screen "101_SDC_PN_Diag128_255" 1280x800, template "SDC"
   on GenerateScreen: SetTag("_intern_BILD_Nr", 101); SetTag("PN_PB\PN\IOSys_ID", 100)
   on ClearScreen: SetTag("_intern_BILD_Nr", 0)
   TextField "OBJECT_674" at 262,49 size 227x27; Text 'ProfiNet-System'
      Visibility <- "PN_PB\IO_Sys_ID"
   Button "Schaltfläche_2" at 240,609 size 107x60; TextOff 'Diagnose PN 101'
      on Press: SetTag("PN_PB\PN\IOSys_ID", 101)
      Visibility <- "PN_PB\IO_Sys_ID"
   Button "Schaltfläche_1" at 240,609 size 107x60; TextOff 'Diagnose PN 100'
      on Press: SetTag("PN_PB\PN\IOSys_ID", 100)
      Visibility <- "PN_PB\IO_Sys_ID"
   Button "Schaltfläche_4" at 573,45 size 359x37; TextOff 'ProfiNet-Teilnehmer 0 - 127'
      on Release: ActivateScreen("100_SDC_PN_Diag0_127", 0)
   GraphicView "OBJECT_496" at 1179,498 size 60x43; Picture "PB_Array_blau_3"
   TextField "OBJECT_497" at 1189,510 size 40x20; Text '1'
   GraphicView "OBJECT_498" at 1179,545 size 60x43; Picture "PB_Array_grün_3"
   TextField "OBJECT_499" at 1189,556 size 40x20; Text '1'
   TextField "OBJECT_500" at 1189,600 size 40x20; Text '1'
   GraphicView "OBJECT_501" at 1179,590 size 60x43; Picture "PB_Array_grün_3"
   TextField "OBJECT_502" at 1189,600 size 40x20; Text '1'
   TextField "OBJECT_504" at 922,505 size 257x31; Text 'Teilnehmer nicht vorhanden'
   TextField "OBJECT_505" at 922,597 size 193x33; Text 'Teilnehmer gestört'
   TextField "OBJECT_506" at 922,552 size 213x33; Text 'Teilnehmer vorhanden'
   TextField "OBJECT_670" at 902,469 size 111x35; Text 'Legende:'
   IOField "OBJECT_675" at 497,50 size 47x29; FormatPattern 999
      ProcessValue <- "PN_PB\IO_Sys_ID"
   TextField "OBJECT_513" at 255,503 size 104x29; Text 'Ort:'
   TextField "OBJECT_514" at 255,533 size 104x31; Text 'Typ:'
   TextField "OBJECT_515" at 255,563 size 131x29; Text 'Bezeichnung:'
   IOField "OBJECT_516" at 399,503 size 167x29; FormatPattern ????????????
      ProcessValue <- "PN_PB\Teiln_Nr_Ort"
   IOField "OBJECT_517" at 399,533 size 156x31; FormatPattern ????????????
      ProcessValue <- "PN_PB\Teiln_Nr_Typ"
   IOField "OBJECT_518" at 399,563 size 253x29; FormatPattern ????????????????????
      ProcessValue <- "PN_PB\Teiln_Nr_Bez"
   IOField "OBJECT_658" at 483,473 size 57x27; FormatPattern 999
      ProcessValue <- "PN_PB\PN\Teiln_Nr"
      Appearance <- "Trigger"
   TextField "OBJECT_679" at 587,473 size 67x25; Text 'Trigger'
      Appearance <- "Trigger"
   GraphicIOField "OBJECT_16" at 749,88 size 60x43; PictureList "PB_Slave_Bit15_3"
      ProcessValue <- "PN_PB\PTMUX_P_TLN129_144"
   GraphicIOField "OBJECT_151" at 813,88 size 60x43; PictureList "PB_Slave_Bit14_3"
      ProcessValue <- "PN_PB\PTMUX_P_TLN129_144"
   GraphicIOField "OBJECT_967" at 874,409 size 60x43; PictureList "PB_Slave_Bit13_3"
      ProcessValue <- "PN_PB\PTMUX_P_TLN241_256"
   GraphicIOField "OBJECT_968" at 1062,409 size 60x43; PictureList "PB_Slave_Bit10_3"
      ProcessValue <- "PN_PB\PTMUX_P_TLN241_256"
   GraphicIOField "OBJECT_969" at 1125,409 size 60x43; PictureList "PB_Slave_Bit9_3"
      ProcessValue <- "PN_PB\PTMUX_P_TLN241_256"
   GraphicIOField "OBJECT_970" at 1187,409 size 60x43; PictureList "PB_Slave_Bit8_3"
      ProcessValue <- "PN_PB\PTMUX_P_TLN241_256"
   GraphicIOField "OBJECT_971" at 999,409 size 60x43; PictureList "PB_Slave_Bit11_3"
      ProcessValue <- "PN_PB\PTMUX_P_TLN241_256"
   GraphicIOField "OBJECT_972" at 811,409 size 60x43; PictureList "PB_Slave_Bit14_3"
      ProcessValue <- "PN_PB\PTMUX_P_TLN241_256"
   GraphicIOField "OBJECT_973" at 937,409 size 60x43; PictureList "PB_Slave_Bit12_3"
      ProcessValue <- "PN_PB\PTMUX_P_TLN241_256"
   GraphicIOField "OBJECT_974" at 749,409 size 60x43; PictureList "PB_Slave_Bit15_3"
      ProcessValue <- "PN_PB\PTMUX_P_TLN241_256"
   GraphicIOField "OBJECT_1030" at 310,409 size 60x43; PictureList "PB_Slave_Bit6_3"
      ProcessValue <- "PN_PB\PTMUX_P_TLN241_256"
   GraphicIOField "OBJECT_1031" at 373,409 size 60x43; PictureList "PB_Slave_Bit5_3"
      ProcessValue <- "PN_PB\PTMUX_P_TLN241_256"
   GraphicIOField "OBJECT_1032" at 435,409 size 60x43; PictureList "PB_Slave_Bit4_3"
      ProcessValue <- "PN_PB\PTMUX_P_TLN241_256"
   GraphicIOField "OBJECT_1033" at 561,409 size 60x43; PictureList "PB_Slave_Bit2_3"
      ProcessValue <- "PN_PB\PTMUX_P_TLN241_256"
   GraphicIOField "OBJECT_1034" at 623,409 size 60x43; PictureList "PB_Slave_Bit1_3"
      ProcessValue <- "PN_PB\PTMUX_P_TLN241_256"
   GraphicIOField "OBJECT_1035" at 686,409 size 60x43; PictureList "PB_Slave_Bit0_3"
      ProcessValue <- "PN_PB\PTMUX_P_TLN241_256"
   GraphicIOField "OBJECT_1036" at 498,409 size 60x43; PictureList "PB_Slave_Bit3_3"
      ProcessValue <- "PN_PB\PTMUX_P_TLN241_256"
   GraphicIOField "OBJECT_1037" at 247,409 size 60x43; PictureList "PB_Slave_Bit7_3"
      ProcessValue <- "PN_PB\PTMUX_P_TLN241_256"
   GraphicIOField "OBJECT_983" at 310,133 size 60x43; PictureList "PB_Slave_Bit6_3"
      ProcessValue <- "PN_PB\PTMUX_P_TLN145_160"
   GraphicIOField "OBJECT_12" at 937,88 size 60x43; PictureList "PB_Slave_Bit12_3"
      ProcessValue <- "PN_PB\PTMUX_P_TLN129_144"
   GraphicIOField "OBJECT_13" at 310,88 size 60x43; PictureList "PB_Slave_Bit6_3"
      ProcessValue <- "PN_PB\PTMUX_P_TLN129_144"
   GraphicIOField "OBJECT_213" at 1062,88 size 60x43; PictureList "PB_Slave_Bit10_3"
      ProcessValue <- "PN_PB\PTMUX_P_TLN129_144"
   GraphicIOField "OBJECT_916" at 1125,88 size 60x43; PictureList "PB_Slave_Bit9_3"
      ProcessValue <- "PN_PB\PTMUX_P_TLN129_144"
   GraphicIOField "OBJECT_917" at 1187,88 size 60x43; PictureList "PB_Slave_Bit8_3"
      ProcessValue <- "PN_PB\PTMUX_P_TLN129_144"
   GraphicIOField "OBJECT_918" at 999,88 size 60x43; PictureList "PB_Slave_Bit11_3"
      ProcessValue <- "PN_PB\PTMUX_P_TLN129_144"
   GraphicIOField "OBJECT_919" at 749,133 size 60x43; PictureList "PB_Slave_Bit15_3"
      ProcessValue <- "PN_PB\PTMUX_P_TLN145_160"
   GraphicIOField "OBJECT_920" at 811,133 size 60x43; PictureList "PB_Slave_Bit14_3"
      ProcessValue <- "PN_PB\PTMUX_P_TLN145_160"
   GraphicIOField "OBJECT_921" at 874,133 size 60x43; PictureList "PB_Slave_Bit13_3"
      ProcessValue <- "PN_PB\PTMUX_P_TLN145_160"
   GraphicIOField "OBJECT_922" at 937,133 size 60x43; PictureList "PB_Slave_Bit12_3"
      ProcessValue <- "PN_PB\PTMUX_P_TLN145_160"
   GraphicIOField "OBJECT_923" at 1062,133 size 60x43; PictureList "PB_Slave_Bit10_3"
      ProcessValue <- "PN_PB\PTMUX_P_TLN145_160"
   GraphicIOField "OBJECT_924" at 1125,133 size 60x43; PictureList "PB_Slave_Bit9_3"
      ProcessValue <- "PN_PB\PTMUX_P_TLN145_160"
   GraphicIOField "OBJECT_925" at 1187,133 size 60x43; PictureList "PB_Slave_Bit8_3"
      ProcessValue <- "PN_PB\PTMUX_P_TLN145_160"
   GraphicIOField "OBJECT_926" at 999,133 size 60x43; PictureList "PB_Slave_Bit11_3"
      ProcessValue <- "PN_PB\PTMUX_P_TLN145_160"
   GraphicIOField "OBJECT_927" at 749,179 size 60x43; PictureList "PB_Slave_Bit15_3"
      ProcessValue <- "PN_PB\PTMUX_P_TLN161_176"
   GraphicIOField "OBJECT_928" at 874,179 size 60x43; PictureList "PB_Slave_Bit13_3"
      ProcessValue <- "PN_PB\PTMUX_P_TLN161_176"
   GraphicIOField "OBJECT_929" at 937,179 size 60x43; PictureList "PB_Slave_Bit12_3"
      ProcessValue <- "PN_PB\PTMUX_P_TLN161_176"
   GraphicIOField "OBJECT_930" at 1062,179 size 60x43; PictureList "PB_Slave_Bit10_3"
      ProcessValue <- "PN_PB\PTMUX_P_TLN161_176"
   GraphicIOField "OBJECT_931" at 1125,179 size 60x43; PictureList "PB_Slave_Bit9_3"
      ProcessValue <- "PN_PB\PTMUX_P_TLN161_176"
   GraphicIOField "OBJECT_932" at 1187,179 size 60x43; PictureList "PB_Slave_Bit8_3"
      ProcessValue <- "PN_PB\PTMUX_P_TLN161_176"
   GraphicIOField "OBJECT_933" at 999,179 size 60x43; PictureList "PB_Slave_Bit11_3"
      ProcessValue <- "PN_PB\PTMUX_P_TLN161_176"
   GraphicIOField "OBJECT_934" at 811,179 size 60x43; PictureList "PB_Slave_Bit14_3"
      ProcessValue <- "PN_PB\PTMUX_P_TLN161_176"
   GraphicIOField "OBJECT_935" at 749,224 size 60x43; PictureList "PB_Slave_Bit15_3"
      ProcessValue <- "PN_PB\PTMUX_P_TLN177_192"
   GraphicIOField "OBJECT_936" at 874,224 size 60x43; PictureList "PB_Slave_Bit13_3"
      ProcessValue <- "PN_PB\PTMUX_P_TLN177_192"
   GraphicIOField "OBJECT_937" at 937,224 size 60x43; PictureList "PB_Slave_Bit12_3"
      ProcessValue <- "PN_PB\PTMUX_P_TLN177_192"
   GraphicIOField "OBJECT_938" at 1062,224 size 60x43; PictureList "PB_Slave_Bit10_3"
      ProcessValue <- "PN_PB\PTMUX_P_TLN177_192"
   GraphicIOField "OBJECT_939" at 1125,224 size 60x43; PictureList "PB_Slave_Bit9_3"
      ProcessValue <- "PN_PB\PTMUX_P_TLN177_192"
   GraphicIOField "OBJECT_940" at 1187,224 size 60x43; PictureList "PB_Slave_Bit8_3"
      ProcessValue <- "PN_PB\PTMUX_P_TLN177_192"
   GraphicIOField "OBJECT_941" at 999,224 size 60x43; PictureList "PB_Slave_Bit11_3"
      ProcessValue <- "PN_PB\PTMUX_P_TLN177_192"
   GraphicIOField "OBJECT_942" at 811,224 size 60x43; PictureList "PB_Slave_Bit14_3"
      ProcessValue <- "PN_PB\PTMUX_P_TLN177_192"
   GraphicIOField "OBJECT_943" at 749,269 size 60x43; PictureList "PB_Slave_Bit15_3"
      ProcessValue <- "PN_PB\PTMUX_P_TLN193_208"
   GraphicIOField "OBJECT_944" at 874,269 size 60x43; PictureList "PB_Slave_Bit13_3"
      ProcessValue <- "PN_PB\PTMUX_P_TLN193_208"
   GraphicIOField "OBJECT_945" at 1062,269 size 60x43; PictureList "PB_Slave_Bit10_3"
      ProcessValue <- "PN_PB\PTMUX_P_TLN193_208"
   GraphicIOField "OBJECT_946" at 1125,269 size 60x43; PictureList "PB_Slave_Bit9_3"
      ProcessValue <- "PN_PB\PTMUX_P_TLN193_208"
   GraphicIOField "OBJECT_947" at 1187,269 size 60x43; PictureList "PB_Slave_Bit8_3"
      ProcessValue <- "PN_PB\PTMUX_P_TLN193_208"
   GraphicIOField "OBJECT_948" at 999,269 size 60x43; PictureList "PB_Slave_Bit11_3"
      ProcessValue <- "PN_PB\PTMUX_P_TLN193_208"
   GraphicIOField "OBJECT_949" at 811,269 size 60x43; PictureList "PB_Slave_Bit14_3"
      ProcessValue <- "PN_PB\PTMUX_P_TLN193_208"
   GraphicIOField "OBJECT_950" at 937,269 size 60x43; PictureList "PB_Slave_Bit12_3"
      ProcessValue <- "PN_PB\PTMUX_P_TLN193_208"
   GraphicIOField "OBJECT_951" at 749,316 size 60x43; PictureList "PB_Slave_Bit15_3"
      ProcessValue <- "PN_PB\PTMUX_P_TLN209_224"
   GraphicIOField "OBJECT_952" at 874,316 size 60x43; PictureList "PB_Slave_Bit13_3"
      ProcessValue <- "PN_PB\PTMUX_P_TLN209_224"
   GraphicIOField "OBJECT_953" at 1062,316 size 60x43; PictureList "PB_Slave_Bit10_3"
      ProcessValue <- "PN_PB\PTMUX_P_TLN209_224"
   GraphicIOField "OBJECT_954" at 1125,316 size 60x43; PictureList "PB_Slave_Bit9_3"
      ProcessValue <- "PN_PB\PTMUX_P_TLN209_224"
   GraphicIOField "OBJECT_955" at 1187,316 size 60x43; PictureList "PB_Slave_Bit8_3"
      ProcessValue <- "PN_PB\PTMUX_P_TLN209_224"
   GraphicIOField "OBJECT_956" at 999,316 size 60x43; PictureList "PB_Slave_Bit11_3"
      ProcessValue <- "PN_PB\PTMUX_P_TLN209_224"
   GraphicIOField "OBJECT_957" at 811,316 size 60x43; PictureList "PB_Slave_Bit14_3"
      ProcessValue <- "PN_PB\PTMUX_P_TLN209_224"
   GraphicIOField "OBJECT_958" at 937,316 size 60x43; PictureList "PB_Slave_Bit12_3"
      ProcessValue <- "PN_PB\PTMUX_P_TLN209_224"
   GraphicIOField "OBJECT_959" at 874,363 size 60x43; PictureList "PB_Slave_Bit13_3"
      ProcessValue <- "PN_PB\PTMUX_P_TLN225_240"
   GraphicIOField "OBJECT_960" at 1062,363 size 60x43; PictureList "PB_Slave_Bit10_3"
      ProcessValue <- "PN_PB\PTMUX_P_TLN225_240"
   GraphicIOField "OBJECT_961" at 1125,363 size 60x43; PictureList "PB_Slave_Bit9_3"
      ProcessValue <- "PN_PB\PTMUX_P_TLN225_240"
   GraphicIOField "OBJECT_962" at 1187,363 size 60x43; PictureList "PB_Slave_Bit8_3"
      ProcessValue <- "PN_PB\PTMUX_P_TLN225_240"
   GraphicIOField "OBJECT_963" at 999,363 size 60x43; PictureList "PB_Slave_Bit11_3"
      ProcessValue <- "PN_PB\PTMUX_P_TLN225_240"
   GraphicIOField "OBJECT_964" at 811,363 size 60x43; PictureList "PB_Slave_Bit14_3"
      ProcessValue <- "PN_PB\PTMUX_P_TLN225_240"
   GraphicIOField "OBJECT_965" at 937,363 size 60x43; PictureList "PB_Slave_Bit12_3"
      ProcessValue <- "PN_PB\PTMUX_P_TLN225_240"
   GraphicIOField "OBJECT_966" at 749,363 size 60x43; PictureList "PB_Slave_Bit15_3"
      ProcessValue <- "PN_PB\PTMUX_P_TLN225_240"
   GraphicIOField "OBJECT_975" at 247,88 size 60x43; PictureList "PB_Slave_Bit7_3"
      ProcessValue <- "PN_PB\PTMUX_P_TLN129_144"
   GraphicIOField "OBJECT_976" at 373,88 size 60x43; PictureList "PB_Slave_Bit5_3"
      ProcessValue <- "PN_PB\PTMUX_P_TLN129_144"
   GraphicIOField "OBJECT_977" at 435,88 size 60x43; PictureList "PB_Slave_Bit4_3"
      ProcessValue <- "PN_PB\PTMUX_P_TLN129_144"
   GraphicIOField "OBJECT_978" at 561,88 size 60x43; PictureList "PB_Slave_Bit2_3"
      ProcessValue <- "PN_PB\PTMUX_P_TLN129_144"
   GraphicIOField "OBJECT_979" at 623,88 size 60x43; PictureList "PB_Slave_Bit1_3"
      ProcessValue <- "PN_PB\PTMUX_P_TLN129_144"
   GraphicIOField "OBJECT_980" at 686,88 size 60x43; PictureList "PB_Slave_Bit0_3"
      ProcessValue <- "PN_PB\PTMUX_P_TLN129_144"
   GraphicIOField "OBJECT_981" at 498,88 size 60x43; PictureList "PB_Slave_Bit3_3"
      ProcessValue <- "PN_PB\PTMUX_P_TLN129_144"
   GraphicIOField "OBJECT_982" at 247,133 size 60x43; PictureList "PB_Slave_Bit7_3"
      ProcessValue <- "PN_PB\PTMUX_P_TLN145_160"
   GraphicIOField "OBJECT_984" at 373,133 size 60x43; PictureList "PB_Slave_Bit5_3"
      ProcessValue <- "PN_PB\PTMUX_P_TLN145_160"
   GraphicIOField "OBJECT_985" at 435,133 size 60x43; PictureList "PB_Slave_Bit4_3"
      ProcessValue <- "PN_PB\PTMUX_P_TLN145_160"
   GraphicIOField "OBJECT_986" at 561,133 size 60x43; PictureList "PB_Slave_Bit2_3"
      ProcessValue <- "PN_PB\PTMUX_P_TLN145_160"
   GraphicIOField "OBJECT_987" at 623,133 size 60x43; PictureList "PB_Slave_Bit1_3"
      ProcessValue <- "PN_PB\PTMUX_P_TLN145_160"
   GraphicIOField "OBJECT_988" at 686,133 size 60x43; PictureList "PB_Slave_Bit0_3"
      ProcessValue <- "PN_PB\PTMUX_P_TLN145_160"
   GraphicIOField "OBJECT_989" at 498,133 size 60x43; PictureList "PB_Slave_Bit3_3"
      ProcessValue <- "PN_PB\PTMUX_P_TLN145_160"
   GraphicIOField "OBJECT_990" at 247,179 size 60x43; PictureList "PB_Slave_Bit7_3"
      ProcessValue <- "PN_PB\PTMUX_P_TLN161_176"
   GraphicIOField "OBJECT_991" at 310,179 size 60x43; PictureList "PB_Slave_Bit6_3"
      ProcessValue <- "PN_PB\PTMUX_P_TLN161_176"
   GraphicIOField "OBJECT_992" at 373,179 size 60x43; PictureList "PB_Slave_Bit5_3"
      ProcessValue <- "PN_PB\PTMUX_P_TLN161_176"
   GraphicIOField "OBJECT_993" at 435,179 size 60x43; PictureList "PB_Slave_Bit4_3"
      ProcessValue <- "PN_PB\PTMUX_P_TLN161_176"
   GraphicIOField "OBJECT_994" at 561,179 size 60x43; PictureList "PB_Slave_Bit2_3"
      ProcessValue <- "PN_PB\PTMUX_P_TLN161_176"
   GraphicIOField "OBJECT_995" at 623,179 size 60x43; PictureList "PB_Slave_Bit1_3"
      ProcessValue <- "PN_PB\PTMUX_P_TLN161_176"
   GraphicIOField "OBJECT_996" at 686,179 size 60x43; PictureList "PB_Slave_Bit0_3"
      ProcessValue <- "PN_PB\PTMUX_P_TLN161_176"
   GraphicIOField "OBJECT_997" at 498,179 size 60x43; PictureList "PB_Slave_Bit3_3"
      ProcessValue <- "PN_PB\PTMUX_P_TLN161_176"
   GraphicIOField "OBJECT_998" at 247,224 size 60x43; PictureList "PB_Slave_Bit7_3"
      ProcessValue <- "PN_PB\PTMUX_P_TLN177_192"
   GraphicIOField "OBJECT_999" at 310,224 size 60x43; PictureList "PB_Slave_Bit6_3"
      ProcessValue <- "PN_PB\PTMUX_P_TLN177_192"
   GraphicIOField "OBJECT_1000" at 375,227 size 60x43; PictureList "PB_Slave_Bit5_3"
      ProcessValue <- "PN_PB\PTMUX_P_TLN177_192"
   GraphicIOField "OBJECT_1001" at 435,224 size 60x43; PictureList "PB_Slave_Bit4_3"
      ProcessValue <- "PN_PB\PTMUX_P_TLN177_192"
   GraphicIOField "OBJECT_1002" at 561,224 size 60x43; PictureList "PB_Slave_Bit2_3"
      ProcessValue <- "PN_PB\PTMUX_P_TLN177_192"
   GraphicIOField "OBJECT_1003" at 623,224 size 60x43; PictureList "PB_Slave_Bit1_3"
      ProcessValue <- "PN_PB\PTMUX_P_TLN177_192"
   GraphicIOField "OBJECT_1004" at 686,224 size 60x43; PictureList "PB_Slave_Bit0_3"
      ProcessValue <- "PN_PB\PTMUX_P_TLN177_192"
   GraphicIOField "OBJECT_1005" at 498,224 size 60x43; PictureList "PB_Slave_Bit3_3"
      ProcessValue <- "PN_PB\PTMUX_P_TLN177_192"
   GraphicIOField "OBJECT_1006" at 247,269 size 60x43; PictureList "PB_Slave_Bit7_3"
      ProcessValue <- "PN_PB\PTMUX_P_TLN193_208"
   GraphicIOField "OBJECT_1007" at 310,269 size 60x43; PictureList "PB_Slave_Bit6_3"
      ProcessValue <- "PN_PB\PTMUX_P_TLN193_208"
   GraphicIOField "OBJECT_1008" at 373,269 size 60x43; PictureList "PB_Slave_Bit5_3"
      ProcessValue <- "PN_PB\PTMUX_P_TLN193_208"
   GraphicIOField "OBJECT_1009" at 435,269 size 60x43; PictureList "PB_Slave_Bit4_3"
      ProcessValue <- "PN_PB\PTMUX_P_TLN193_208"
   GraphicIOField "OBJECT_1010" at 561,269 size 60x43; PictureList "PB_Slave_Bit2_3"
      ProcessValue <- "PN_PB\PTMUX_P_TLN193_208"
   GraphicIOField "OBJECT_1011" at 623,269 size 60x43; PictureList "PB_Slave_Bit1_3"
      ProcessValue <- "PN_PB\PTMUX_P_TLN193_208"
   GraphicIOField "OBJECT_1012" at 686,269 size 60x43; PictureList "PB_Slave_Bit0_3"
      ProcessValue <- "PN_PB\PTMUX_P_TLN193_208"
   GraphicIOField "OBJECT_1013" at 498,269 size 60x43; PictureList "PB_Slave_Bit3_3"
      ProcessValue <- "PN_PB\PTMUX_P_TLN193_208"
   GraphicIOField "OBJECT_1014" at 247,316 size 60x43; PictureList "PB_Slave_Bit7_3"
      ProcessValue <- "PN_PB\PTMUX_P_TLN209_224"
   GraphicIOField "OBJECT_1015" at 310,316 size 60x43; PictureList "PB_Slave_Bit6_3"
      ProcessValue <- "PN_PB\PTMUX_P_TLN209_224"
   GraphicIOField "OBJECT_1016" at 373,316 size 60x43; PictureList "PB_Slave_Bit5_3"
      ProcessValue <- "PN_PB\PTMUX_P_TLN209_224"
   GraphicIOField "OBJECT_1017" at 435,316 size 60x43; PictureList "PB_Slave_Bit4_3"
      ProcessValue <- "PN_PB\PTMUX_P_TLN209_224"
   GraphicIOField "OBJECT_1018" at 561,316 size 60x43; PictureList "PB_Slave_Bit2_3"
      ProcessValue <- "PN_PB\PTMUX_P_TLN209_224"
   GraphicIOField "OBJECT_1019" at 623,316 size 60x43; PictureList "PB_Slave_Bit1_3"
      ProcessValue <- "PN_PB\PTMUX_P_TLN209_224"
   GraphicIOField "OBJECT_1020" at 686,316 size 60x43; PictureList "PB_Slave_Bit0_3"
      ProcessValue <- "PN_PB\PTMUX_P_TLN209_224"
   GraphicIOField "OBJECT_1021" at 498,316 size 60x43; PictureList "PB_Slave_Bit3_3"
      ProcessValue <- "PN_PB\PTMUX_P_TLN209_224"
   GraphicIOField "OBJECT_1022" at 247,363 size 60x43; PictureList "PB_Slave_Bit7_3"
      ProcessValue <- "PN_PB\PTMUX_P_TLN225_240"
   GraphicIOField "OBJECT_1023" at 310,363 size 60x43; PictureList "PB_Slave_Bit6_3"
      ProcessValue <- "PN_PB\PTMUX_P_TLN225_240"
   GraphicIOField "OBJECT_1024" at 373,363 size 60x43; PictureList "PB_Slave_Bit5_3"
      ProcessValue <- "PN_PB\PTMUX_P_TLN225_240"
   GraphicIOField "OBJECT_1025" at 435,363 size 60x43; PictureList "PB_Slave_Bit4_3"
      ProcessValue <- "PN_PB\PTMUX_P_TLN225_240"
   GraphicIOField "OBJECT_1026" at 561,363 size 60x43; PictureList "PB_Slave_Bit2_3"
      ProcessValue <- "PN_PB\PTMUX_P_TLN225_240"
   GraphicIOField "OBJECT_1027" at 623,363 size 60x43; PictureList "PB_Slave_Bit1_3"
      ProcessValue <- "PN_PB\PTMUX_P_TLN225_240"
   GraphicIOField "OBJECT_1028" at 686,363 size 60x43; PictureList "PB_Slave_Bit0_3"
      ProcessValue <- "PN_PB\PTMUX_P_TLN225_240"
   GraphicIOField "OBJECT_1029" at 498,363 size 60x43; PictureList "PB_Slave_Bit3_3"
      ProcessValue <- "PN_PB\PTMUX_P_TLN225_240"
   GraphicIOField "OBJECT_14" at 874,88 size 60x43; PictureList "PB_Slave_Bit13_3"
      ProcessValue <- "PN_PB\PTMUX_P_TLN129_144"
   TextField "OBJECT_508" at 255,473 size 227x27; Text 'Profibus-Teilnehmer:'
      Visibility <- "PN_PB\IO_Sys_ID"
   TextField "OBJECT_306" at 1198,99 size 40x20; Text '128'
      Appearance <- "PN_PB\PTMUX_F_TLN129_144"
   TextField "OBJECT_340" at 1137,99 size 40x20; Text '129'
      Appearance <- "PN_PB\PTMUX_F_TLN129_144"
   TextField "OBJECT_372" at 1073,99 size 40x20; Text '130'
      Appearance <- "PN_PB\PTMUX_F_TLN129_144"
   TextField "OBJECT_374" at 1010,99 size 40x20; Text '131'
      Appearance <- "PN_PB\PTMUX_F_TLN129_144"
   TextField "OBJECT_408" at 949,99 size 40x20; Text '132'
      Appearance <- "PN_PB\PTMUX_F_TLN129_144"
   TextField "OBJECT_410" at 822,99 size 40x20; Text '134'
      Appearance <- "PN_PB\PTMUX_F_TLN129_144"
   TextField "OBJECT_443" at 759,99 size 40x20; Text '135'
      Appearance <- "PN_PB\PTMUX_F_TLN129_144"
   TextField "OBJECT_509" at 1135,144 size 40x20; Text '145'
      Appearance <- "PN_PB\PTMUX_F_TLN145_160"
   TextField "OBJECT_510" at 1073,144 size 40x20; Text '146'
      Appearance <- "PN_PB\PTMUX_F_TLN145_160"
   TextField "OBJECT_512" at 1010,144 size 40x20; Text '147'
      Appearance <- "PN_PB\PTMUX_F_TLN145_160"
   TextField "OBJECT_677" at 947,144 size 40x20; Text '148'
      Appearance <- "PN_PB\PTMUX_F_TLN145_160"
   TextField "OBJECT_678" at 885,144 size 40x20; Text '149'
      Appearance <- "PN_PB\PTMUX_F_TLN145_160"
   TextField "OBJECT_680" at 822,144 size 40x20; Text '150'
      Appearance <- "PN_PB\PTMUX_F_TLN145_160"
   TextField "OBJECT_681" at 759,144 size 40x20; Text '151'
      Appearance <- "PN_PB\PTMUX_F_TLN145_160"
   TextField "OBJECT_682" at 1198,144 size 40x20; Text '144'
      Appearance <- "PN_PB\PTMUX_F_TLN145_160"
   TextField "OBJECT_691" at 1198,189 size 40x20; Text '160'
      Appearance <- "PN_PB\PTMUX_F_TLN161_176"
   TextField "OBJECT_692" at 1135,189 size 40x20; Text '161'
      Appearance <- "PN_PB\PTMUX_F_TLN161_176"
   TextField "OBJECT_693" at 1073,189 size 40x20; Text '162'
      Appearance <- "PN_PB\PTMUX_F_TLN161_176"
   TextField "OBJECT_694" at 1010,189 size 40x20; Text '163'
      Appearance <- "PN_PB\PTMUX_F_TLN161_176"
   TextField "OBJECT_695" at 947,189 size 40x20; Text '164'
      Appearance <- "PN_PB\PTMUX_F_TLN161_176"
   TextField "OBJECT_696" at 885,189 size 40x20; Text '165'
      Appearance <- "PN_PB\PTMUX_F_TLN161_176"
   TextField "OBJECT_697" at 759,189 size 40x20; Text '167'
      Appearance <- "PN_PB\PTMUX_F_TLN161_176"
   TextField "OBJECT_699" at 822,189 size 40x20; Text '166'
      Appearance <- "PN_PB\PTMUX_F_TLN161_176"
   TextField "OBJECT_708" at 1198,235 size 40x20; Text '176'
      Appearance <- "PN_PB\PTMUX_F_TLN177_192"
   TextField "OBJECT_709" at 1135,235 size 40x20; Text '177'
      Appearance <- "PN_PB\PTMUX_F_TLN177_192"
   TextField "OBJECT_710" at 1073,235 size 40x20; Text '178'
      Appearance <- "PN_PB\PTMUX_F_TLN177_192"
   TextField "OBJECT_711" at 947,235 size 40x20; Text '180'
      Appearance <- "PN_PB\PTMUX_F_TLN177_192"
   TextField "OBJECT_712" at 885,235 size 40x20; Text '181'
      Appearance <- "PN_PB\PTMUX_F_TLN177_192"
   TextField "OBJECT_713" at 759,235 size 40x20; Text '183'
      Appearance <- "PN_PB\PTMUX_F_TLN177_192"
   TextField "OBJECT_715" at 822,235 size 40x20; Text '182'
      Appearance <- "PN_PB\PTMUX_F_TLN177_192"
   TextField "OBJECT_716" at 1010,235 size 40x20; Text '179'
      Appearance <- "PN_PB\PTMUX_F_TLN177_192"
   TextField "OBJECT_724" at 1198,281 size 40x20; Text '192'
      Appearance <- "PN_PB\PTMUX_F_TLN193_208"
   TextField "OBJECT_725" at 1135,281 size 40x20; Text '193'
      Appearance <- "PN_PB\PTMUX_F_TLN193_208"
   TextField "OBJECT_726" at 1073,281 size 40x20; Text '194'
      Appearance <- "PN_PB\PTMUX_F_TLN193_208"
   TextField "OBJECT_727" at 885,281 size 40x20; Text '197'
      Appearance <- "PN_PB\PTMUX_F_TLN193_208"
   TextField "OBJECT_728" at 759,281 size 40x20; Text '199'
      Appearance <- "PN_PB\PTMUX_F_TLN193_208"
   TextField "OBJECT_730" at 822,281 size 40x20; Text '198'
      Appearance <- "PN_PB\PTMUX_F_TLN193_208"
   TextField "OBJECT_731" at 1010,281 size 40x20; Text '195'
      Appearance <- "PN_PB\PTMUX_F_TLN193_208"
   TextField "OBJECT_733" at 947,281 size 40x20; Text '196'
      Appearance <- "PN_PB\PTMUX_F_TLN193_208"
   TextField "OBJECT_741" at 1198,328 size 40x20; Text '208'
      Appearance <- "PN_PB\PTMUX_F_TLN209_224"
   TextField "OBJECT_742" at 1135,328 size 40x20; Text '209'
      Appearance <- "PN_PB\PTMUX_F_TLN209_224"
   TextField "OBJECT_743" at 1073,328 size 40x20; Text '210'
      Appearance <- "PN_PB\PTMUX_F_TLN209_224"
   TextField "OBJECT_744" at 885,328 size 40x20; Text '213'
      Appearance <- "PN_PB\PTMUX_F_TLN209_224"
   TextField "OBJECT_746" at 822,328 size 40x20; Text '214'
      Appearance <- "PN_PB\PTMUX_F_TLN209_224"
   TextField "OBJECT_747" at 1010,328 size 40x20; Text '211'
      Appearance <- "PN_PB\PTMUX_F_TLN209_224"
   TextField "OBJECT_749" at 947,328 size 40x20; Text '212'
      Appearance <- "PN_PB\PTMUX_F_TLN209_224"
   TextField "OBJECT_750" at 759,328 size 40x20; Text '215'
      Appearance <- "PN_PB\PTMUX_F_TLN209_224"
   TextField "OBJECT_757" at 1198,375 size 40x20; Text '224'
      Appearance <- "PN_PB\PTMUX_F_TLN225_240"
   TextField "OBJECT_758" at 1135,375 size 40x20; Text '225'
      Appearance <- "PN_PB\PTMUX_F_TLN225_240"
   TextField "OBJECT_759" at 1073,375 size 40x20; Text '226'
      Appearance <- "PN_PB\PTMUX_F_TLN225_240"
   TextField "OBJECT_760" at 885,375 size 40x20; Text '229'
      Appearance <- "PN_PB\PTMUX_F_TLN225_240"
   TextField "OBJECT_762" at 822,375 size 40x20; Text '230'
      Appearance <- "PN_PB\PTMUX_F_TLN225_240"
   TextField "OBJECT_763" at 1010,375 size 40x20; Text '227'
      Appearance <- "PN_PB\PTMUX_F_TLN225_240"
   TextField "OBJECT_765" at 947,375 size 40x20; Text '228'
      Appearance <- "PN_PB\PTMUX_F_TLN225_240"
   TextField "OBJECT_767" at 759,375 size 40x20; Text '231'
      Appearance <- "PN_PB\PTMUX_F_TLN225_240"
   TextField "OBJECT_774" at 1198,420 size 40x20; Text '240'
      Appearance <- "PN_PB\PTMUX_F_TLN241_256"
   TextField "OBJECT_775" at 1135,420 size 40x20; Text '241'
      Appearance <- "PN_PB\PTMUX_F_TLN241_256"
   TextField "OBJECT_776" at 1073,420 size 40x20; Text '242'
      Appearance <- "PN_PB\PTMUX_F_TLN241_256"
   TextField "OBJECT_777" at 885,420 size 40x20; Text '245'
      Appearance <- "PN_PB\PTMUX_F_TLN241_256"
   TextField "OBJECT_779" at 822,420 size 40x20; Text '246'
      Appearance <- "PN_PB\PTMUX_F_TLN241_256"
   TextField "OBJECT_780" at 1010,420 size 40x20; Text '243'
      Appearance <- "PN_PB\PTMUX_F_TLN241_256"
   TextField "OBJECT_782" at 947,420 size 40x20; Text '244'
      Appearance <- "PN_PB\PTMUX_F_TLN241_256"
   TextField "OBJECT_784" at 759,420 size 40x20; Text '247'
      Appearance <- "PN_PB\PTMUX_F_TLN241_256"
   TextField "OBJECT_787" at 697,99 size 40x20; Text '136'
      Appearance <- "PN_PB\PTMUX_F_TLN129_144"
   TextField "OBJECT_789" at 634,99 size 40x20; Text '137'
      Appearance <- "PN_PB\PTMUX_F_TLN129_144"
   TextField "OBJECT_790" at 571,99 size 40x20; Text '138'
      Appearance <- "PN_PB\PTMUX_F_TLN129_144"
   TextField "OBJECT_791" at 509,99 size 40x20; Text '139'
      Appearance <- "PN_PB\PTMUX_F_TLN129_144"
   TextField "OBJECT_792" at 446,99 size 40x20; Text '140'
      Appearance <- "PN_PB\PTMUX_F_TLN129_144"
   TextField "OBJECT_793" at 383,99 size 40x20; Text '141'
      Appearance <- "PN_PB\PTMUX_F_TLN129_144"
   TextField "OBJECT_794" at 321,99 size 40x20; Text '142'
      Appearance <- "PN_PB\PTMUX_F_TLN129_144"
   TextField "OBJECT_795" at 258,99 size 40x20; Text '143'
      Appearance <- "PN_PB\PTMUX_F_TLN129_144"
   TextField "OBJECT_804" at 697,144 size 40x20; Text '152'
      Appearance <- "PN_PB\PTMUX_F_TLN145_160"
   TextField "OBJECT_806" at 634,144 size 40x20; Text '153'
      Appearance <- "PN_PB\PTMUX_F_TLN145_160"
   TextField "OBJECT_807" at 571,144 size 40x20; Text '154'
      Appearance <- "PN_PB\PTMUX_F_TLN145_160"
   TextField "OBJECT_808" at 509,144 size 40x20; Text '155'
      Appearance <- "PN_PB\PTMUX_F_TLN145_160"
   TextField "OBJECT_809" at 446,144 size 40x20; Text '156'
      Appearance <- "PN_PB\PTMUX_F_TLN145_160"
   TextField "OBJECT_810" at 383,144 size 40x20; Text '157'
      Appearance <- "PN_PB\PTMUX_F_TLN145_160"
   TextField "OBJECT_811" at 321,144 size 40x20; Text '158'
      Appearance <- "PN_PB\PTMUX_F_TLN145_160"
   TextField "OBJECT_812" at 258,144 size 40x20; Text '159'
      Appearance <- "PN_PB\PTMUX_F_TLN145_160"
   TextField "OBJECT_821" at 697,189 size 40x20; Text '168'
      Appearance <- "PN_PB\PTMUX_F_TLN161_176"
   TextField "OBJECT_823" at 634,189 size 40x20; Text '169'
      Appearance <- "PN_PB\PTMUX_F_TLN161_176"
   TextField "OBJECT_824" at 571,189 size 40x20; Text '170'
      Appearance <- "PN_PB\PTMUX_F_TLN161_176"
   TextField "OBJECT_825" at 509,189 size 40x20; Text '171'
      Appearance <- "PN_PB\PTMUX_F_TLN161_176"
   TextField "OBJECT_826" at 446,189 size 40x20; Text '172'
      Appearance <- "PN_PB\PTMUX_F_TLN161_176"
   TextField "OBJECT_827" at 383,189 size 40x20; Text '173'
      Appearance <- "PN_PB\PTMUX_F_TLN161_176"
   TextField "OBJECT_828" at 321,189 size 40x20; Text '174'
      Appearance <- "PN_PB\PTMUX_F_TLN161_176"
   TextField "OBJECT_829" at 258,189 size 40x20; Text '175'
      Appearance <- "PN_PB\PTMUX_F_TLN161_176"
   TextField "OBJECT_838" at 697,235 size 40x20; Text '184'
      Appearance <- "PN_PB\PTMUX_F_TLN177_192"
   TextField "OBJECT_840" at 634,235 size 40x20; Text '185'
      Appearance <- "PN_PB\PTMUX_F_TLN177_192"
   TextField "OBJECT_841" at 571,235 size 40x20; Text '186'
      Appearance <- "PN_PB\PTMUX_F_TLN177_192"
   TextField "OBJECT_842" at 509,235 size 40x20; Text '187'
      Appearance <- "PN_PB\PTMUX_F_TLN177_192"
   TextField "OBJECT_843" at 446,235 size 40x20; Text '188'
      Appearance <- "PN_PB\PTMUX_F_TLN177_192"
   TextField "OBJECT_844" at 383,235 size 40x20; Text '189'
      Appearance <- "PN_PB\PTMUX_F_TLN177_192"
   TextField "OBJECT_845" at 321,235 size 40x20; Text '190'
      Appearance <- "PN_PB\PTMUX_F_TLN177_192"
   TextField "OBJECT_846" at 258,235 size 40x20; Text '191'
      Appearance <- "PN_PB\PTMUX_F_TLN177_192"
   TextField "OBJECT_855" at 697,281 size 40x20; Text '200'
      Appearance <- "PN_PB\PTMUX_F_TLN193_208"
   TextField "OBJECT_857" at 634,281 size 40x20; Text '201'
      Appearance <- "PN_PB\PTMUX_F_TLN193_208"
   TextField "OBJECT_858" at 571,281 size 40x20; Text '202'
      Appearance <- "PN_PB\PTMUX_F_TLN193_208"
   TextField "OBJECT_859" at 509,281 size 40x20; Text '203'
      Appearance <- "PN_PB\PTMUX_F_TLN193_208"
   TextField "OBJECT_860" at 446,281 size 40x20; Text '204'
      Appearance <- "PN_PB\PTMUX_F_TLN193_208"
   TextField "OBJECT_861" at 383,281 size 40x20; Text '205'
      Appearance <- "PN_PB\PTMUX_F_TLN193_208"
   TextField "OBJECT_862" at 321,281 size 40x20; Text '206'
      Appearance <- "PN_PB\PTMUX_F_TLN193_208"
   TextField "OBJECT_863" at 258,281 size 40x20; Text '207'
      Appearance <- "PN_PB\PTMUX_F_TLN193_208"
   TextField "OBJECT_872" at 697,328 size 40x20; Text '216'
      Appearance <- "PN_PB\PTMUX_F_TLN209_224"
   TextField "OBJECT_874" at 634,328 size 40x20; Text '217'
      Appearance <- "PN_PB\PTMUX_F_TLN209_224"
   TextField "OBJECT_875" at 571,328 size 40x20; Text '218'
      Appearance <- "PN_PB\PTMUX_F_TLN209_224"
   TextField "OBJECT_876" at 509,328 size 40x20; Text '219'
      Appearance <- "PN_PB\PTMUX_F_TLN209_224"
   TextField "OBJECT_877" at 446,328 size 40x20; Text '220'
      Appearance <- "PN_PB\PTMUX_F_TLN209_224"
   TextField "OBJECT_878" at 383,328 size 40x20; Text '221'
      Appearance <- "PN_PB\PTMUX_F_TLN209_224"
   TextField "OBJECT_879" at 321,328 size 40x20; Text '222'
      Appearance <- "PN_PB\PTMUX_F_TLN209_224"
   TextField "OBJECT_880" at 258,328 size 40x20; Text '223'
      Appearance <- "PN_PB\PTMUX_F_TLN209_224"
   TextField "OBJECT_889" at 697,375 size 40x20; Text '232'
      Appearance <- "PN_PB\PTMUX_F_TLN225_240"
   TextField "OBJECT_891" at 634,375 size 40x20; Text '233'
      Appearance <- "PN_PB\PTMUX_F_TLN225_240"
   TextField "OBJECT_892" at 571,375 size 40x20; Text '234'
      Appearance <- "PN_PB\PTMUX_F_TLN225_240"
   TextField "OBJECT_893" at 509,375 size 40x20; Text '235'
      Appearance <- "PN_PB\PTMUX_F_TLN225_240"
   TextField "OBJECT_894" at 446,375 size 40x20; Text '236'
      Appearance <- "PN_PB\PTMUX_F_TLN225_240"
   TextField "OBJECT_895" at 383,375 size 40x20; Text '237'
      Appearance <- "PN_PB\PTMUX_F_TLN225_240"
   TextField "OBJECT_896" at 321,375 size 40x20; Text '238'